// TIA Portal project "XSFW_TIA32701_A6" (V15.1) (continued)
REGION Network 6: en ciclo
   RUNG wire#powerrail
      Contact( "iPls_Marcha" )
      wire#w1
      S_SR(operand := "En_ciclo", r1 := wire#w2)
      wire#w3
      R_Coil( "Comandos".marcha_panel )
   END_RUNG
   RUNG wire#powerrail
      Contact( "Comandos".marcha_panel )
   END_RUNG wire#w1
   RUNG wire#powerrail
      I_Contact( "iPls_Parada" )
   END_RUNG wire#w2
   RUNG wire#powerrail
      Contact( "iSns_Solapa_Abierta" )
   END_RUNG wire#w2
   RUNG wire#powerrail
      Contact( "Comandos".parada_panel )
   END_RUNG wire#w2
   RUNG wire#powerrail
      I_Contact( "iGmt_rolos_Ent" )
   END_RUNG wire#w2
   RUNG wire#powerrail
      I_Contact( "iGmt_cin_later" )
   END_RUNG wire#w2
   RUNG wire#powerrail
      I_Contact( "Circuito_Seguridad" )
   END_RUNG wire#w2
   RUNG wire#powerrail
      Contact( "Falla_rol_entra" )
   END_RUNG wire#w2
   RUNG wire#powerrail
      I_Contact( "Marcha_Linea" )
   END_RUNG wire#w2
   RUNG wire#powerrail
      P_Contact(operand := "Alarma Activa", bit := "Tag_2")
   END_RUNG wire#w2
   RUNG wire#w3
      Not()
      R_Coil( "Comandos".parada_panel )
   END_RUNG
   // the same network as SCL:
   #_w1 := "Alarma Activa" AND NOT "Tag_2";   // rising edge of "Alarma Activa"
   "Tag_2" := "Alarma Activa";
   IF "iPls_Marcha" OR "Comandos".marcha_panel THEN
       "En_ciclo" := TRUE;   // SR flip-flop
   END_IF;
   IF NOT "iPls_Parada" OR "iSns_Solapa_Abierta" OR "Comandos".parada_panel OR NOT "iGmt_rolos_Ent" OR NOT "iGmt_cin_later" OR NOT "Circuito_Seguridad" OR "Falla_rol_entra" OR NOT "Marcha_Linea" OR #_w1 THEN
       "En_ciclo" := FALSE;
   END_IF;
   IF "En_ciclo" THEN "Comandos".marcha_panel := FALSE; END_IF;
   IF NOT "En_ciclo" THEN "Comandos".parada_panel := FALSE; END_IF;
END_REGION

REGION Network 7: SALIDA A0.5 - falla presente
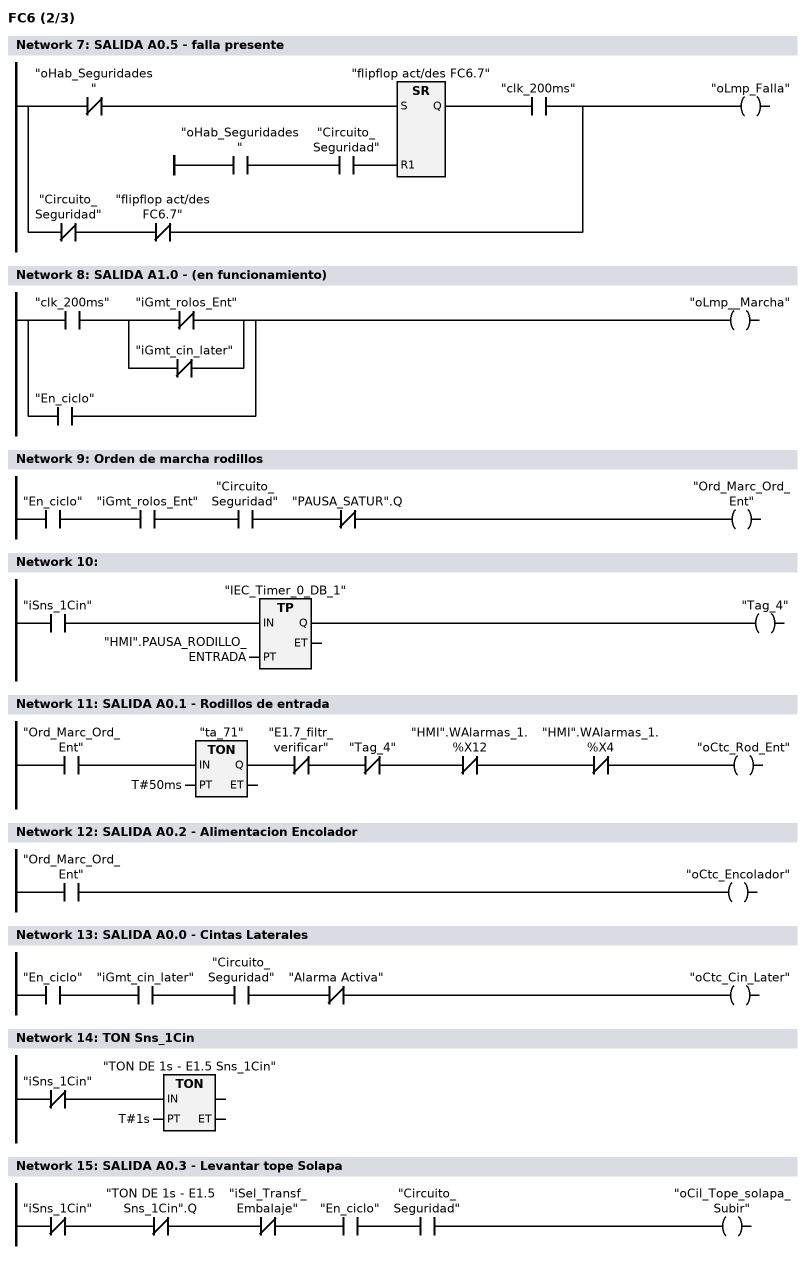
   RUNG wire#powerrail
      I_Contact( "oHab_Seguridades" )
      S_SR(operand := "flipflop act/des FC6.7", r1 := wire#w1)
      Contact( "clk_200ms" )
      wire#w2
      Coil( "oLmp_Falla" )
   END_RUNG
   RUNG wire#powerrail
      Contact( "oHab_Seguridades" )
      Contact( "Circuito_Seguridad" )
   END_RUNG wire#w1
   RUNG wire#powerrail
      I_Contact( "Circuito_Seguridad" )
      I_Contact( "flipflop act/des FC6.7" )
   END_RUNG wire#w2
   // the same network as SCL:
   IF NOT "oHab_Seguridades" THEN
       "flipflop act/des FC6.7" := TRUE;   // SR flip-flop
   END_IF;
   IF "oHab_Seguridades" AND "Circuito_Seguridad" THEN "flipflop act/des FC6.7" := FALSE; END_IF;
   "oLmp_Falla" := ("flipflop act/des FC6.7" AND "clk_200ms") OR (NOT "Circuito_Seguridad" AND NOT "flipflop act/des FC6.7");
END_REGION

REGION Network 8: SALIDA A1.0 - (en funcionamiento)
   RUNG wire#powerrail
      Contact( "clk_200ms" )
      wire#w1
      I_Contact( "iGmt_rolos_Ent" )
      wire#w2
      Coil( "oLmp__Marcha" )
   END_RUNG
   RUNG wire#w1
      I_Contact( "iGmt_cin_later" )
   END_RUNG wire#w2
   RUNG wire#powerrail
      Contact( "En_ciclo" )
   END_RUNG wire#w2
   // the same network as SCL:
   "oLmp__Marcha" := ("clk_200ms" AND (NOT "iGmt_rolos_Ent" OR NOT "iGmt_cin_later")) OR "En_ciclo";
END_REGION

REGION Network 9: Orden de marcha rodillos
   RUNG wire#powerrail
      Contact( "En_ciclo" )
      Contact( "iGmt_rolos_Ent" )
      Contact( "Circuito_Seguridad" )
      I_Contact( "PAUSA_SATUR".Q )
      Coil( "Ord_Marc_Ord_Ent" )
   END_RUNG
   // the same network as SCL:
   "Ord_Marc_Ord_Ent" := "En_ciclo" AND "iGmt_rolos_Ent" AND "Circuito_Seguridad" AND NOT "PAUSA_SATUR".Q;
END_REGION

REGION Network 10
   "IEC_Timer_0_DB_1".TP(IN := "iSns_1Cin", PT := "HMI".PAUSA_RODILLO_ENTRADA);
   "Tag_4" := "IEC_Timer_0_DB_1".Q;
END_REGION

REGION Network 11: SALIDA A0.1 - Rodillos de entrada
   "ta_71".TON(IN := "Ord_Marc_Ord_Ent", PT := T#50ms);
   "oCtc_Rod_Ent" := "ta_71".Q AND NOT "E1.7_filtr_verificar" AND NOT "Tag_4" AND NOT "HMI".WAlarmas_1.%X12 AND NOT "HMI".WAlarmas_1.%X4;
END_REGION

REGION Network 12: SALIDA A0.2 - Alimentacion Encolador
   RUNG wire#powerrail
      Contact( "Ord_Marc_Ord_Ent" )
      Coil( "oCtc_Encolador" )
   END_RUNG
   // the same network as SCL:
   "oCtc_Encolador" := "Ord_Marc_Ord_Ent";
END_REGION

REGION Network 13: SALIDA A0.0 - Cintas Laterales
   RUNG wire#powerrail
      Contact( "En_ciclo" )
      Contact( "iGmt_cin_later" )
      Contact( "Circuito_Seguridad" )
      I_Contact( "Alarma Activa" )
      Coil( "oCtc_Cin_Later" )
   END_RUNG
   // the same network as SCL:
   "oCtc_Cin_Later" := "En_ciclo" AND "iGmt_cin_later" AND "Circuito_Seguridad" AND NOT "Alarma Activa";
END_REGION

REGION Network 14: TON Sns_1Cin
   "TON DE 1s - E1.5 Sns_1Cin".TON(IN := NOT "iSns_1Cin", PT := T#1s);
END_REGION

REGION Network 15: SALIDA A0.3 - Levantar tope Solapa
   RUNG wire#powerrail
      I_Contact( "iSns_1Cin" )
      I_Contact( "TON DE 1s - E1.5 Sns_1Cin".Q )
      I_Contact( "iSel_Transf_Embalaje" )
      Contact( "En_ciclo" )
      Contact( "Circuito_Seguridad" )
      Coil( "oCil_Tope_solapa_Subir" )
   END_RUNG
   // the same network as SCL:
   "oCil_Tope_solapa_Subir" := NOT "iSns_1Cin" AND NOT "TON DE 1s - E1.5 Sns_1Cin".Q AND NOT "iSel_Transf_Embalaje" AND "En_ciclo" AND "Circuito_Seguridad";
END_REGION

REGION Network 16: Orden bajar tope solapa trtasera
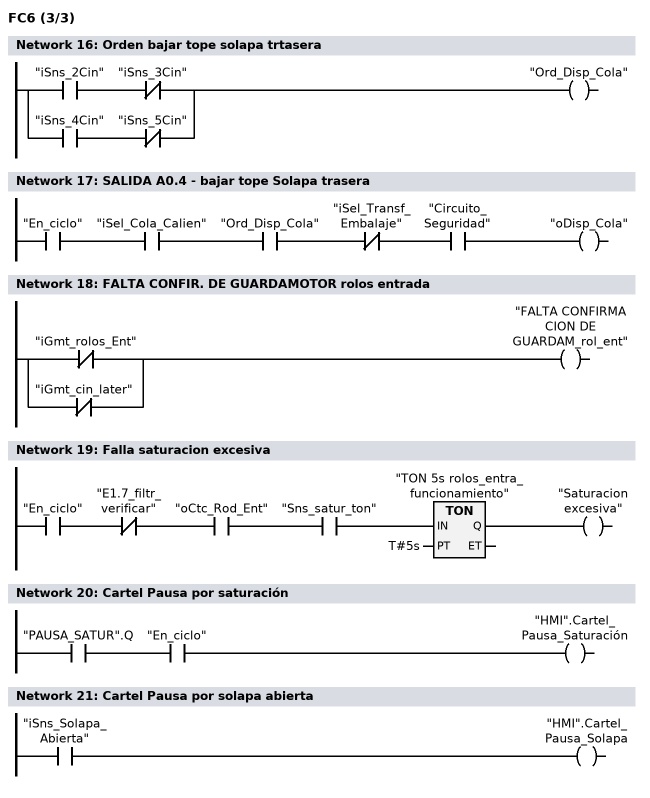
   RUNG wire#powerrail
      Contact( "iSns_2Cin" )
      I_Contact( "iSns_3Cin" )
      wire#w1
      Coil( "Ord_Disp_Cola" )
   END_RUNG
   RUNG wire#powerrail
      Contact( "iSns_4Cin" )
      I_Contact( "iSns_5Cin" )
   END_RUNG wire#w1
   // the same network as SCL:
   "Ord_Disp_Cola" := ("iSns_2Cin" AND NOT "iSns_3Cin") OR ("iSns_4Cin" AND NOT "iSns_5Cin");
END_REGION

REGION Network 17: SALIDA A0.4 - bajar tope Solapa trasera
   RUNG wire#powerrail
      Contact( "En_ciclo" )
      Contact( "iSel_Cola_Calien" )
      Contact( "Ord_Disp_Cola" )
      I_Contact( "iSel_Transf_Embalaje" )
      Contact( "Circuito_Seguridad" )
      Coil( "oDisp_Cola" )
   END_RUNG
   // the same network as SCL:
   "oDisp_Cola" := "En_ciclo" AND "iSel_Cola_Calien" AND "Ord_Disp_Cola" AND NOT "iSel_Transf_Embalaje" AND "Circuito_Seguridad";
END_REGION

REGION Network 18: FALTA CONFIR. DE GUARDAMOTOR rolos entrada
   RUNG wire#powerrail
      I_Contact( "iGmt_rolos_Ent" )
      wire#w1
      Coil( "FALTA CONFIRMACION DE GUARDAM_rol_ent" )
   END_RUNG
   RUNG wire#powerrail
      I_Contact( "iGmt_cin_later" )
   END_RUNG wire#w1
   // the same network as SCL:
   "FALTA CONFIRMACION DE GUARDAM_rol_ent" := NOT "iGmt_rolos_Ent" OR NOT "iGmt_cin_later";
END_REGION

REGION Network 19: Falla saturacion excesiva
   "TON 5s rolos_entra_ funcionamiento".TON(IN := "En_ciclo" AND NOT "E1.7_filtr_verificar" AND "oCtc_Rod_Ent" AND "Sns_satur_ton",
                           PT := T#5s);
   "Saturacion excesiva" := "TON 5s rolos_entra_ funcionamiento".Q;
END_REGION

REGION Network 20: Cartel Pausa por saturación
   RUNG wire#powerrail
      Contact( "PAUSA_SATUR".Q )
      Contact( "En_ciclo" )
      Coil( "HMI".Cartel_Pausa_Saturación )
   END_RUNG
   // the same network as SCL:
   "HMI".Cartel_Pausa_Saturación := "PAUSA_SATUR".Q AND "En_ciclo";
END_REGION

REGION Network 21: Cartel Pausa por solapa abierta
   RUNG wire#powerrail
      Contact( "iSns_Solapa_Abierta" )
      Coil( "HMI".Cartel_Pausa_Solapa )
   END_RUNG
   // the same network as SCL:
   "HMI".Cartel_Pausa_Solapa := "iSns_Solapa_Abierta";
END_REGION
END_FUNCTION

FUNCTION "FC10" : Void   // FC10, LAD
{ S7_Optimized_Access := 'TRUE' }
VERSION : 0.1
BEGIN

REGION Network 1: SALIDA A1.1 - Habilitacion de seguridades
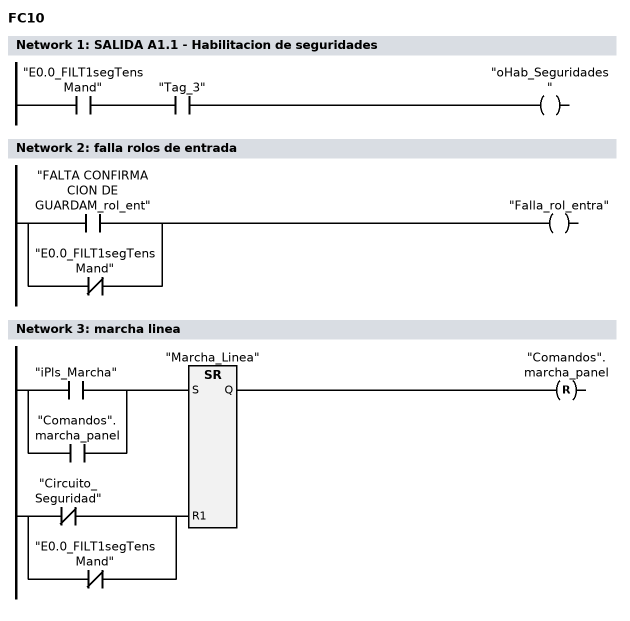
   RUNG wire#powerrail
      Contact( "E0.0_FILT1segTensMand" )
      Contact( "Tag_3" )
      Coil( "oHab_Seguridades" )
   END_RUNG
   // the same network as SCL:
   "oHab_Seguridades" := "E0.0_FILT1segTensMand" AND "Tag_3";
END_REGION

REGION Network 2: falla rolos de entrada
   RUNG wire#powerrail
      Contact( "FALTA CONFIRMACION DE GUARDAM_rol_ent" )
      wire#w1
      Coil( "Falla_rol_entra" )
   END_RUNG
   RUNG wire#powerrail
      I_Contact( "E0.0_FILT1segTensMand" )
   END_RUNG wire#w1
   // the same network as SCL:
   "Falla_rol_entra" := "FALTA CONFIRMACION DE GUARDAM_rol_ent" OR NOT "E0.0_FILT1segTensMand";
END_REGION

REGION Network 3: marcha linea
   RUNG wire#powerrail
      Contact( "iPls_Marcha" )
      wire#w1
      S_SR(operand := "Marcha_Linea", r1 := wire#w2)
      R_Coil( "Comandos".marcha_panel )
   END_RUNG
   RUNG wire#powerrail
      Contact( "Comandos".marcha_panel )
   END_RUNG wire#w1
   RUNG wire#powerrail
      I_Contact( "Circuito_Seguridad" )
   END_RUNG wire#w2
   RUNG wire#powerrail
      I_Contact( "E0.0_FILT1segTensMand" )
   END_RUNG wire#w2
   // the same network as SCL:
   IF "iPls_Marcha" OR "Comandos".marcha_panel THEN
       "Marcha_Linea" := TRUE;   // SR flip-flop
   END_IF;
   IF NOT "Circuito_Seguridad" OR NOT "E0.0_FILT1segTensMand" THEN "Marcha_Linea" := FALSE; END_IF;
   IF "Marcha_Linea" THEN "Comandos".marcha_panel := FALSE; END_IF;
END_REGION
END_FUNCTION

ORGANIZATION_BLOCK "OB1"   // OB1, LAD, ProgramCycle
TITLE = "Main Program Sweep (Cycle)"
{ S7_Optimized_Access := 'TRUE' }
VERSION : 0.1
   VAR_INPUT
      Initial_Call : Bool;   // Initial call of this OB
      Remanence : Bool;   // =True, if remanent data are available
   END_VAR
BEGIN

REGION Network 1: Marcas de Sistema
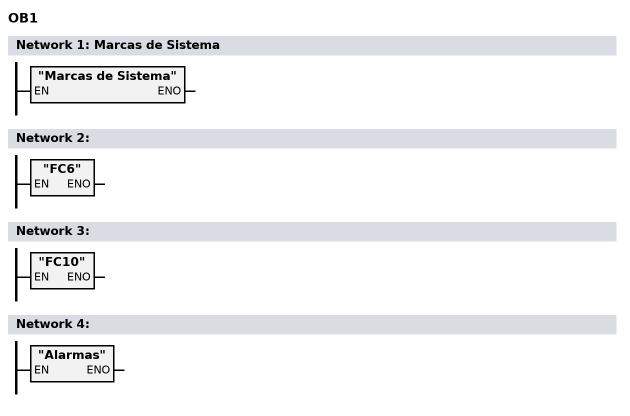
   RUNG wire#powerrail
      "Marcas de Sistema"()
   END_RUNG
   // the same network as SCL:
   "Marcas de Sistema"();
END_REGION

REGION Network 2
   RUNG wire#powerrail
      "FC6"()
   END_RUNG
   // the same network as SCL:
   "FC6"();
END_REGION

REGION Network 3
   RUNG wire#powerrail
      "FC10"()
   END_RUNG
   // the same network as SCL:
   "FC10"();
END_REGION

REGION Network 4
   RUNG wire#powerrail
      "Alarmas"()
   END_RUNG
   // the same network as SCL:
   "Alarmas"();
END_REGION
END_ORGANIZATION_BLOCK

(* ===== HMI "HMI_RT_1" =====
system functions are stored by id; their names below are inferred from use
connection "HMI_Conexión_1": ETHERNET, SMART_S7_1200_OMS

HMI tags "Tabla de variables estándar"
   "DB1_D_5" : Word = PLC DB1.D_5 AT %DB1.DBW10, 1 s
   "comandos_marcha_panel" : Bool = PLC Comandos.marcha_panel, 1 s
   "HMI_Tiem_Satur" : Time = PLC HMI.Tiem_Satur, 1 s
   "HMI_Tiem_saturPan" : Time = PLC HMI.Tiem_Satur, 1 s
   "comandos_parada_panel" : Bool = PLC Comandos.parada_panel, 1 s
   "WAlarmas_1" : Word = PLC HMI.WAlarmas_1 AT %DB1.DBW0, 1 s
   "HMI_RESET" : Bool = PLC HMI.RESET, 1 s
   "Tension_Mando" : Bool = PLC iTension_Mando AT %I0.0, 1 s
   "Guard_cin_later" : Bool = PLC iGmt_cin_later AT %I0.3, 1 s
   "Guard_rolos_Ent" : Bool = PLC iGmt_rolos_Ent AT %I0.4, 1 s
   "Parad_Emerg" : Bool = PLC iParad_Emerg AT %I0.1, 1 s
   "Puerta_1" : Bool = PLC iSns_Puerta_1 AT %I2.0, 1 s
   "Puerta_2" : Bool = PLC iSns_Puerta_2 AT %I2.1, 1 s
   "Puerta_3" : Bool = PLC iSns_Puerta_3 AT %I2.2, 1 s
   "Puerta_4" : Bool = PLC iSns_Puerta_4 AT %I2.3, 1 s
   "En_ciclo" : Bool = PLC En_ciclo AT %M161.0, 1 s
   "Alarma Activa" : Bool = PLC "Alarma Activa" AT %M10.0, 1 s
   "Pul_Marcha" : Bool = PLC iPls_Marcha AT %I0.5, 1 s
   "Puls_parada" : Bool = PLC iPls_Parada AT %I0.6, 1 s
   "Selec_Transf_Embalaje" : Bool = PLC iSel_Transf_Embalaje AT %I0.7, 1 s
   "Selec_Cola_Calien" : Bool = PLC iSel_Cola_Calien AT %I1.0, 1 s
   "Sns_2Cin" : Bool = PLC iSns_2Cin AT %I1.1, 1 s
   "Sns_3Cin" : Bool = PLC iSns_3Cin AT %I1.2, 1 s
   "Sns_4Cin" : Bool = PLC iSns_4Cin AT %I1.3, 1 s
   "Sns_5Cin" : Bool = PLC iSns_5Cin AT %I1.4, 1 s
   "Sns_1Cin" : Bool = PLC iSns_1Cin AT %I1.5, 1 s
   "Sns_Satur" : Bool = PLC iSns_Satur AT %I1.6, 1 s
   "RELEVAR_SIEMP_LLEGA_1" : Bool = PLC RELEVAR_SIEMP_LLEGA_1 AT %I1.7, 1 s
   "SOLAPA ABIERTA" : Bool = PLC iSns_Solapa_Abierta AT %I2.4, 1 s
   "Saturacion excesiva" : Bool = PLC "Saturacion excesiva" AT %M160.5, 1 s
   "PAUSA_SATUR_Q" : Bool = PLC PAUSA_SATUR.Q, 1 s
   "iReserva I0.2" : Bool = PLC "iReserva RESET I0.2" AT %I0.2, 1 s
   "iReserva I2.5" : Bool = PLC "iReserva I2.5" AT %I2.5, 1 s
   "iReserva I2.6" : Bool = PLC "iReserva I2.6" AT %I2.6, 1 s
   "iReserva I2.7" : Bool = PLC "iReserva I2.7" AT %I2.7, 1 s
   "oCtc_Cin_Later" : Bool = PLC oCtc_Cin_Later AT %Q0.0, 1 s
   "oCtc_Rod_Ent" : Bool = PLC oCtc_Rod_Ent AT %Q0.1, 1 s
   "oCtc_Encolador" : Bool = PLC oCtc_Encolador AT %Q0.2, 1 s
   "oCil_Tope_solapa_Subir" : Bool = PLC oCil_Tope_solapa_Subir AT %Q0.3, 1 s
   "oCil_Tope_solapa_Bajar" : Bool = PLC oDisp_Cola AT %Q0.4, 1 s
   "oLmp_Falla" : Bool = PLC oLmp_Falla AT %Q0.5, 1 s
   "oLmp__Marcha" : Bool = PLC oLmp__Marcha AT %Q1.0, 1 s
   "oHab_Seguridades" : Bool = PLC oHab_Seguridades AT %Q1.1, 1 s
   "oReserva A1.2" : Bool = PLC "oReserva A1.2" AT %Q1.2, 1 s
   "oReserva A1.3" : Bool = PLC "oReserva A1.3" AT %Q1.3, 1 s
   "oReserva A1.4" : Bool = PLC "oReserva A1.4" AT %Q1.4, 1 s
   "oReserva A1.5" : Bool = PLC "oReserva A1.5" AT %Q1.5, 1 s
   "oReserva A1.6" : Bool = PLC "oReserva A1.6" AT %Q1.6, 1 s
   "oReserva A1.7" : Bool = PLC "oReserva A1.7" AT %Q1.7, 1 s
   "oReserva A2.0" : Bool = PLC "oReserva A2.0" AT %Q2.0, 1 s
   "oReserva A2.1" : Bool = PLC "oReserva A2.1" AT %Q2.1, 1 s
   "oReserva A2.2" : Bool = PLC "oReserva A2.2" AT %Q2.2, 1 s
   "oReserva A2.3" : Bool = PLC "oReserva A2.3" AT %Q2.3, 1 s
   "oReserva A2.4" : Bool = PLC "oReserva A2.4" AT %Q2.4, 1 s
   "oReserva A2.5" : Bool = PLC "oReserva A2.5" AT %Q2.5, 1 s
   "oReserva A2.6" : Bool = PLC "oReserva A2.6" AT %Q2.6, 1 s
   "oReserva A2.7" : Bool = PLC "oReserva A2.7" AT %Q2.7, 1 s
   "HMI_Cartel_Pausa_Saturación" : Bool = PLC HMI.Cartel_Pausa_Saturación, 1 s
   "HMI_Cartel_Pausa_Solapa" : Bool = PLC HMI.Cartel_Pausa_Solapa, 1 s
   "HMI_PAUSA_RODILLO_ENTRADA" : Time = PLC HMI.PAUSA_RODILLO_ENTRADA, 1 s
   "Temporizadores_Tiempo1" : Time = PLC Temporizadores.Tiempo1, 1 s

discrete alarms
   1: 'FALLA EN SEGURIDAD', class Warnings, trigger "WAlarmas_1" bit 0
   2: 'GUARDAMOTOR ROLOS ENTRADA', class Warnings, trigger "WAlarmas_1" bit 1
   3: 'GUARDAMOTOR CINTAS LATERALES', class Warnings, trigger "WAlarmas_1" bit 2
   4: 'ALIMENTACION ENCOLADOR', class Warnings, trigger "WAlarmas_1" bit 3
   5: 'TIEMPO DE SATURCION EXCEDIDA', class Warnings, trigger "WAlarmas_1" bit 4
   6: 'PARADA DE EMERGENCIA ACTIVA', class Warnings, trigger "WAlarmas_1" bit 5
   7: 'PUERTA 1', class Warnings, trigger "WAlarmas_1" bit 6
   8: 'PUERTA 2', class Warnings, trigger "WAlarmas_1" bit 7
   9: 'PUERTA 3', class Warnings, trigger "WAlarmas_1" bit 8
   10: 'PUERTA 4', class Warnings, trigger "WAlarmas_1" bit 9
   11: 'SOLAPA ABIERTA', class Warnings, trigger "WAlarmas_1" bit 10
   12: 'Falta tension 24VDC en E0.0', class Warnings, trigger "WAlarmas_1" bit 11
   13: 'Tiempo excesivo de Cola', class Warnings, trigger "WAlarmas_1" bit 12

screen "INICIO" 800x480, template "Plantilla_1"
   GraphicView "Visor de gráficos_1" at 0,0 size 800x432; Picture "XING_MOD317_A0"
   Button "Botón_1" at 223,47 size 137x57; TextOff 'MARCHA'
      on Click: SetBit("comandos_marcha_panel")
   Button "Botón_2" at 371,47 size 137x57; TextOff 'PARADA'
      on Click: SetBit("comandos_parada_panel")
   Button "Botón_3" at 642,47 size 137x57; TextOff 'RESET'
      on Click: SetBit("HMI_RESET")
   Rectangle "Rectángulo_1" at 117,371 size 108x36
      Appearance <- "Puerta_1"
   TextField "Campo de texto_1" at 135,376 size 75x23; Text 'Puerta 1'
   Rectangle "Rectángulo_2" at 229,371 size 108x36
      Appearance <- "Puerta_2"
   TextField "Campo de texto_2" at 247,376 size 75x23; Text 'Puerta 2'
   Rectangle "Rectángulo_3" at 341,371 size 108x36
      Appearance <- "Puerta_3"
   TextField "Campo de texto_3" at 359,376 size 75x23; Text 'Puerta 3'
   Rectangle "Rectángulo_4" at 453,371 size 108x36
      Appearance <- "Puerta_4"
   TextField "Campo de texto_4" at 471,376 size 75x23; Text 'Puerta 4'
   Rectangle "Rectángulo_5" at 565,371 size 108x36
      Appearance <- "Parad_Emerg"
   TextField "Campo de texto_5" at 567,376 size 100x23; Text 'Emergencia'
   Button "Botón_4" at 223,47 size 137x57; TextOff 'MARCHA'
      on Click: SetBit("comandos_marcha_panel")
      Visibility <- "En_ciclo"
   Button "Botón_5" at 371,47 size 137x57; TextOff 'PARADA'
      on Click: SetBit("comandos_parada_panel")
      Visibility <- "En_ciclo"
   Button "Botón_6" at 642,47 size 137x57; TextOff 'RESET'
      on Click: SetBit("HMI_RESET")
      Visibility <- "Alarma Activa"
   Rectangle "Rectángulo_6" at 12,150 size 142x68
      Visibility <- "HMI_Cartel_Pausa_Solapa"
   TextField "Campo de texto_6" at 16,162 size 134x42; Text 'Parada por Solapa Abierta'
      Visibility <- "SOLAPA ABIERTA"
   Rectangle "Rectángulo_7" at 12,150 size 142x68
      Visibility <- "HMI_Cartel_Pausa_Saturación"
   TextField "Campo de texto_7" at 30,163 size 100x42; Text 'Pausa por Saturación'
      Visibility <- "HMI_Cartel_Pausa_Saturación"

screen "TIEMPOS" 800x480, template "Plantilla_1"
   GraphicView "Visor de gráficos_1" at 0,0 size 800x433; Picture "XING_MOD317_A0"
   IOField "Campo ES_2" at 28,192 size 116x32; FormatPattern 99999; Unit  segs.
      ProcessValue <- "HMI_Tiem_saturPan"
   TextField "Campo de texto_1" at 20,139 size 129x42; Text 'Tiempo Pausa por Saturación'
   IOField "Campo ES_1" at 604,106 size 116x32; FormatPattern 99999; Unit  segs.
      ProcessValue <- "HMI_PAUSA_RODILLO_ENTRADA"
   TextField "Campo de texto_2" at 596,53 size 120x42; Text 'Tiempo Pausa Entre Cajas'
   IOField "Campo ES_3" at 332,82 size 116x32; FormatPattern 99999; Unit  segs.
      ProcessValue <- "Temporizadores_Tiempo1"
   TextField "Campo de texto_3" at 312,35 size 156x42; Text 'Alarma de Disparo de Cola'

screen "ALARMAS" 800x480, template "Plantilla_1"
   AlarmView "Visor de avisos_1" at 23,56 size 756x347

Template "Plantilla_1" 800x480
   Button "Botón_2" at 480,432 size 161x48; TextOff 'Salidas'
      on Click: ActivateScreen("SALIDAS 1/2", 0)
   Button "Botón_3" at 320,432 size 161x48; TextOff 'Tiempos'
      on Click: ActivateScreen("TIEMPOS", 0)
   Button "Botón_4" at 160,432 size 161x48; TextOff 'Entradas'
      on Click: ActivateScreen("ENTRADAS 1/2", 0)
   Button "Botón_6" at 0,432 size 161x48; TextOff 'Principal'
      on Click: ActivateScreen("INICIO", 0)
   Button "Botón_1" at 639,432 size 161x48; TextOff 'Alarmas'
      on Click: ActivateScreen("ALARMAS", 0)
   DateTimeField "Plantilla_Campo de fecha y hora_1" at 596,2 size 197x24
   GraphicView "Plantilla_Visor de gráficos_1" at 9,2 size 76x24; Picture "eProC Logo Paneles Parte B"

screen "ENTRADAS 1/2" 800x480, template "Plantilla_1"
   Circle "Círculo_1" at 21,38 size 46x46
      Appearance <- "Tension_Mando"
   TextField "Campo de texto_1" at 24,49 size 43x23; Text 'E0.0'
   Circle "Círculo_2" at 21,38 size 46x46
      Appearance <- "Tension_Mando"
   TextField "Campo de texto_2" at 24,49 size 43x23; Text 'E0.0'
   Circle "Círculo_3" at 21,86 size 46x46
      Appearance <- "Parad_Emerg"
   TextField "Campo de texto_3" at 24,97 size 43x23; Text 'E0.1'
   Circle "Círculo_4" at 21,134 size 46x46
      Appearance <- "iReserva I0.2"
   TextField "Campo de texto_4" at 24,145 size 43x23; Text 'E0.2'
   Circle "Círculo_5" at 21,182 size 46x46
      Appearance <- "Guard_cin_later"
   TextField "Campo de texto_5" at 24,193 size 43x23; Text 'E0.3'
   Circle "Círculo_6" at 21,230 size 46x46
      Appearance <- "Guard_rolos_Ent"
   TextField "Campo de texto_6" at 24,241 size 43x23; Text 'E0.4'
   Circle "Círculo_7" at 21,278 size 46x46
      Appearance <- "Pul_Marcha"
   TextField "Campo de texto_7" at 24,289 size 43x23; Text 'E0.5'
   Circle "Círculo_8" at 21,326 size 46x46
      Appearance <- "Puls_parada"
   TextField "Campo de texto_8" at 24,337 size 43x23; Text 'E0.6'
   Circle "Círculo_25" at 21,374 size 46x46
      Appearance <- "Selec_Transf_Embalaje"
   TextField "Campo de texto_25" at 24,385 size 43x23; Text 'E0.7'
   TextField "Campo de texto_9" at 72,49 size 154x23; Text 'Tensión de mando'
   TextField "Campo de texto_10" at 72,97 size 188x23; Text 'Parada de emergencia'
   TextField "Campo de texto_11" at 72,193 size 246x23; Text 'Guardamotor Cintas laterales'
   TextField "Campo de texto_12" at 72,241 size 232x23; Text 'Guardamotor Rolos entrada'
   TextField "Campo de texto_14" at 72,289 size 165x23; Text 'Pulsador de Marcha'
   TextField "Campo de texto_15" at 72,337 size 164x23; Text 'Pulsador de Parada'
   TextField "Campo de texto_16" at 72,385 size 213x23; Text 'Selectora tranf. embalaje'
   Circle "Círculo_9" at 357,38 size 46x46
      Appearance <- "Tension_Mando"
   TextField "Campo de texto_13" at 360,49 size 43x23; Text 'E0.0'
   Circle "Círculo_10" at 357,38 size 46x46
      Appearance <- "Selec_Cola_Calien"
   TextField "Campo de texto_17" at 360,49 size 43x23; Text 'E1.0'
   Circle "Círculo_11" at 357,86 size 46x46
      Appearance <- "Sns_2Cin"
   TextField "Campo de texto_18" at 360,97 size 43x23; Text 'E1.1'
   Circle "Círculo_12" at 357,134 size 46x46
      Appearance <- "Sns_3Cin"
   TextField "Campo de texto_19" at 360,145 size 43x23; Text 'E1.2'
   Circle "Círculo_13" at 357,182 size 46x46
      Appearance <- "Sns_4Cin"
   TextField "Campo de texto_20" at 360,193 size 43x23; Text 'E1.3'
   Circle "Círculo_14" at 357,230 size 46x46
      Appearance <- "Sns_5Cin"
   TextField "Campo de texto_21" at 360,241 size 43x23; Text 'E1.4'
   Circle "Círculo_15" at 357,278 size 46x46
      Appearance <- "Sns_1Cin"
   TextField "Campo de texto_22" at 360,289 size 43x23; Text 'E1.5'
   Circle "Círculo_16" at 357,326 size 46x46
      Appearance <- "Sns_Satur"
   TextField "Campo de texto_23" at 360,337 size 43x23; Text 'E1.6'
   Circle "Círculo_17" at 357,374 size 46x46
      Appearance <- "RELEVAR_SIEMP_LLEGA_1"
   TextField "Campo de texto_24" at 360,385 size 43x23; Text 'E1.7'
   TextField "Campo de texto_26" at 408,49 size 190x23; Text 'Selectora cola caliente'
   TextField "Campo de texto_27" at 408,97 size 123x23; Text 'Sensor 2 Cinta'
   TextField "Campo de texto_28" at 408,193 size 123x23; Text 'Sensor 4 Cinta'
   TextField "Campo de texto_29" at 408,241 size 123x23; Text 'Sensor 5 Cinta'
   TextField "Campo de texto_30" at 408,289 size 123x23; Text 'Sensor 1 Cinta'
   TextField "Campo de texto_31" at 408,337 size 175x23; Text 'Sensor de saturación'
   TextField "Campo de texto_33" at 408,145 size 123x23; Text 'Sensor 3 Cinta'
   TextField "Campo de texto_32" at 72,145 size 71x23; Text 'Reserva'
   TextField "Campo de texto_34" at 408,385 size 71x23; Text 'Reserva'
   Button "Botón_1" at 716,104 size 73x49; TextOff 'PÁG 2'
      on Click: ActivateScreen("ENTRADAS 2/2", 0)
   Button "Botón_2" at 716,48 size 73x49; TextOff 'PÁG 1'
      on Click: ActivateScreen("ENTRADAS 1/2", 0)
   Button "Botón_3" at 716,48 size 73x49; TextOff 'PÁG 1'
      on Click: ActivateScreen("ENTRADAS 1/2", 0)

screen "ENTRADAS 2/2" 800x480, template "Plantilla_1"
   Circle "Círculo_1" at 21,38 size 46x46
      Appearance <- "Tension_Mando"
   TextField "Campo de texto_1" at 24,49 size 43x23; Text 'E0.0'
   Circle "Círculo_2" at 21,38 size 46x46
      Appearance <- "Puerta_1"
   TextField "Campo de texto_2" at 24,49 size 43x23; Text 'E2.0'
   Circle "Círculo_3" at 21,86 size 46x46
      Appearance <- "Puerta_2"
   TextField "Campo de texto_3" at 24,97 size 43x23; Text 'E2.1'
   Circle "Círculo_4" at 21,134 size 46x46
      Appearance <- "Puerta_3"
   TextField "Campo de texto_4" at 24,145 size 43x23; Text 'E2.2'
   Circle "Círculo_5" at 21,182 size 46x46
      Appearance <- "Puerta_4"
   TextField "Campo de texto_5" at 24,193 size 43x23; Text 'E2.3'
   Circle "Círculo_6" at 21,230 size 46x46
      Appearance <- "SOLAPA ABIERTA"
   TextField "Campo de texto_6" at 24,241 size 43x23; Text 'E2.4'
   Circle "Círculo_7" at 21,278 size 46x46
      Appearance <- "iReserva I2.5"
   TextField "Campo de texto_7" at 24,289 size 43x23; Text 'E2.5'
   Circle "Círculo_8" at 21,326 size 46x46
      Appearance <- "iReserva I2.6"
   TextField "Campo de texto_8" at 24,337 size 43x23; Text 'E2.6'
   Circle "Círculo_25" at 21,374 size 46x46
      Appearance <- "iReserva I2.7"
   TextField "Campo de texto_25" at 24,385 size 43x23; Text 'E2.7'
   TextField "Campo de texto_9" at 72,49 size 75x23; Text 'Puerta 1'
   TextField "Campo de texto_10" at 72,97 size 75x23; Text 'Puerta 2'
   TextField "Campo de texto_12" at 72,241 size 209x23; Text 'Sensor de Solapa abierta'
   TextField "Campo de texto_11" at 72,145 size 75x23; Text 'Puerta 3'
   TextField "Campo de texto_32" at 72,193 size 75x23; Text 'Puerta 4'
   TextField "Campo de texto_14" at 72,289 size 71x23; Text 'Reserva'
   TextField "Campo de texto_15" at 72,337 size 71x23; Text 'Reserva'
   TextField "Campo de texto_16" at 72,385 size 71x23; Text 'Reserva'
   Button "Botón_1" at 716,104 size 73x49; TextOff 'PÁG 2'
      on Click: ActivateScreen("ENTRADAS 2/2", 0)
   Button "Botón_2" at 716,48 size 73x49; TextOff 'PÁG 1'
      on Click: ActivateScreen("ENTRADAS 1/2", 0)
   Button "Botón_4" at 716,104 size 73x49; TextOff 'PÁG 2'
      on Click: ActivateScreen("ENTRADAS 2/2", 0)

screen "SALIDAS 2/2" 800x480, template "Plantilla_1"
   Circle "Círculo_9" at 21,38 size 46x46
      Appearance <- "Tension_Mando"
   TextField "Campo de texto_13" at 24,49 size 43x23; Text 'E0.0'
   Circle "Círculo_10" at 21,38 size 46x46
      Appearance <- "oReserva A2.0"
   TextField "Campo de texto_17" at 22,49 size 43x23; Text 'A2.0'
   Circle "Círculo_11" at 21,86 size 46x46
      Appearance <- "oReserva A2.1"
   TextField "Campo de texto_18" at 22,97 size 43x23; Text 'A2.1'
   Circle "Círculo_12" at 21,134 size 46x46
      Appearance <- "oReserva A2.2"
   TextField "Campo de texto_19" at 22,145 size 43x23; Text 'A2.2'
   Circle "Círculo_13" at 21,182 size 46x46
      Appearance <- "oReserva A2.3"
   TextField "Campo de texto_20" at 22,193 size 43x23; Text 'A2.3'
   Circle "Círculo_14" at 21,230 size 46x46
      Appearance <- "oReserva A2.4"
   TextField "Campo de texto_21" at 22,241 size 43x23; Text 'A2.4'
   Circle "Círculo_15" at 21,278 size 46x46
      Appearance <- "oReserva A2.5"
   TextField "Campo de texto_22" at 22,289 size 43x23; Text 'A2.5'
   TextField "Campo de texto_26" at 72,49 size 71x23; Text 'Reserva'
   Circle "Círculo_1" at 21,326 size 46x46
      Appearance <- "oReserva A2.6"
   TextField "Campo de texto_23" at 22,337 size 43x23; Text 'A2.6'
   Circle "Círculo_16" at 21,374 size 46x46
      Appearance <- "oReserva A2.7"
   TextField "Campo de texto_31" at 22,385 size 43x23; Text 'A2.7'
   TextField "Campo de texto_1" at 72,97 size 71x23; Text 'Reserva'
   TextField "Campo de texto_2" at 72,145 size 71x23; Text 'Reserva'
   TextField "Campo de texto_3" at 72,193 size 71x23; Text 'Reserva'
   TextField "Campo de texto_4" at 72,241 size 71x23; Text 'Reserva'
   TextField "Campo de texto_5" at 72,289 size 71x23; Text 'Reserva'
   TextField "Campo de texto_6" at 72,337 size 71x23; Text 'Reserva'
   TextField "Campo de texto_7" at 72,385 size 71x23; Text 'Reserva'
   Button "Botón_1" at 716,104 size 73x49; TextOff 'PÁG 2'
      on Click: ActivateScreen("SALIDAS 2/2", 0)
   Button "Botón_4" at 716,104 size 73x49; TextOff 'PÁG 2'
      on Click: ActivateScreen("SALIDAS 2/2", 0)
   Button "Botón_2" at 716,48 size 73x49; TextOff 'PÁG 1'
      on Click: ActivateScreen("SALIDAS 1/2", 0)

screen "SALIDAS 1/2" 800x480, template "Plantilla_1"
   Circle "Círculo_9" at 21,38 size 46x46
      Appearance <- "Tension_Mando"
   TextField "Campo de texto_13" at 24,49 size 43x23; Text 'E0.0'
   Circle "Círculo_10" at 21,38 size 46x46
      Appearance <- "oCtc_Cin_Later"
   TextField "Campo de texto_17" at 22,49 size 43x23; Text 'A0.0'
   Circle "Círculo_11" at 21,86 size 46x46
      Appearance <- "oCtc_Rod_Ent"
   TextField "Campo de texto_18" at 22,97 size 43x23; Text 'A0.1'
   Circle "Círculo_12" at 21,134 size 46x46
      Appearance <- "oCtc_Encolador"
   TextField "Campo de texto_19" at 22,145 size 43x23; Text 'A0.2'
   Circle "Círculo_13" at 21,182 size 46x46
      Appearance <- "oCil_Tope_solapa_Subir"
   TextField "Campo de texto_20" at 22,193 size 43x23; Text 'A0.3'
   Circle "Círculo_14" at 21,230 size 46x46
      Appearance <- "oCil_Tope_solapa_Bajar"
   TextField "Campo de texto_21" at 22,241 size 43x23; Text 'A0.4'
   Circle "Círculo_15" at 21,278 size 46x46
      Appearance <- "oLmp_Falla"
   TextField "Campo de texto_22" at 22,289 size 43x23; Text 'A0.5'
   TextField "Campo de texto_26" at 72,49 size 197x23; Text 'Marcha Cintas laterales'
   TextField "Campo de texto_27" at 72,97 size 203x23; Text 'Marcha Rodillos entrada'
   TextField "Campo de texto_28" at 72,193 size 147x23; Text 'Subir tope solapa'
   TextField "Campo de texto_29" at 72,241 size 149x23; Text 'Bajar tope solapa'
   TextField "Campo de texto_30" at 72,289 size 204x23; Text 'Indicador luminoso Falla'
   TextField "Campo de texto_33" at 72,145 size 173x23; Text 'Encendido encolador'
   Circle "Círculo_2" at 357,38 size 46x46
      Appearance <- "Tension_Mando"
   TextField "Campo de texto_1" at 360,49 size 43x23; Text 'E0.0'
   Circle "Círculo_3" at 357,38 size 46x46
      Appearance <- "oLmp__Marcha"
   TextField "Campo de texto_2" at 358,49 size 43x23; Text 'A1.0'
   Circle "Círculo_4" at 357,86 size 46x46
      Appearance <- "oHab_Seguridades"
   TextField "Campo de texto_3" at 358,97 size 43x23; Text 'A1.1'
   Circle "Círculo_5" at 357,134 size 46x46
      Appearance <- "oReserva A1.2"
   TextField "Campo de texto_4" at 358,145 size 43x23; Text 'A1.2'
   Circle "Círculo_6" at 357,182 size 46x46
      Appearance <- "oReserva A1.3"
   TextField "Campo de texto_5" at 358,193 size 43x23; Text 'A1.3'
   Circle "Círculo_7" at 357,230 size 46x46
      Appearance <- "oReserva A1.4"
   TextField "Campo de texto_6" at 358,241 size 43x23; Text 'A1.4'
   Circle "Círculo_8" at 357,278 size 46x46
      Appearance <- "oReserva A1.5"
   TextField "Campo de texto_7" at 358,289 size 43x23; Text 'A1.5'
   Circle "Círculo_18" at 357,326 size 46x46
      Appearance <- "oReserva A1.6"
   TextField "Campo de texto_8" at 358,337 size 43x23; Text 'A1.6'
   Circle "Círculo_19" at 357,374 size 46x46
      Appearance <- "oReserva A1.7"
   TextField "Campo de texto_9" at 358,385 size 43x23; Text 'A1.7'
   TextField "Campo de texto_10" at 408,49 size 224x23; Text 'Indicador luminoso Marcha'
   TextField "Campo de texto_11" at 408,97 size 230x23; Text 'Habilitación de seguridades'
   TextField "Campo de texto_12" at 408,193 size 71x23; Text 'Reserva'
   TextField "Campo de texto_14" at 408,241 size 71x23; Text 'Reserva'
   TextField "Campo de texto_15" at 408,289 size 71x23; Text 'Reserva'
   TextField "Campo de texto_16" at 408,337 size 71x23; Text 'Reserva'
   TextField "Campo de texto_25" at 408,145 size 71x23; Text 'Reserva'
   TextField "Campo de texto_32" at 408,385 size 71x23; Text 'Reserva'
   Button "Botón_1" at 716,104 size 73x49; TextOff 'PÁG 2'
      on Click: ActivateScreen("SALIDAS 2/2", 0)
   Button "Botón_2" at 716,48 size 73x49; TextOff 'PÁG 1'
      on Click: ActivateScreen("SALIDAS 1/2", 0)
   Button "Botón_3" at 716,48 size 73x49; TextOff 'PÁG 1'
      on Click: ActivateScreen("SALIDAS 1/2", 0)
*)